   864: 'Spare_Fault_864', class No Acknowledgement, trigger "DB302_HMI_Faults_Carrier13_Faults_1" bit 15
   865: 'Carrier 13 Motion Off Fault', class No Acknowledgement, trigger "DB302_HMI_Faults_Carrier13_Faults_2" bit 0
   866: 'Carrier 13 Motion On Fault', class No Acknowledgement, trigger "DB302_HMI_Faults_Carrier13_Faults_2" bit 1
   867: 'Carrier 13 Spacing Fault', class No Acknowledgement, trigger "DB302_HMI_Faults_Carrier13_Faults_2" bit 2
   868: 'Carrier 13 Duplicate Carrier Number Fault', class No Acknowledgement, trigger "DB302_HMI_Faults_Carrier13_Faults_2" bit 3
   869: 'Spare_Fault_869', class No Acknowledgement, trigger "DB302_HMI_Faults_Carrier13_Faults_2" bit 4
   870: 'Spare_Fault_870', class No Acknowledgement, trigger "DB302_HMI_Faults_Carrier13_Faults_2" bit 5
   871: 'Spare_Fault_871', class No Acknowledgement, trigger "DB302_HMI_Faults_Carrier13_Faults_2" bit 6
   872: 'Spare_Fault_872', class No Acknowledgement, trigger "DB302_HMI_Faults_Carrier13_Faults_2" bit 7
   873: 'Spare_Fault_873', class No Acknowledgement, trigger "DB302_HMI_Faults_Carrier13_Faults_2" bit 8
   874: 'Spare_Fault_874', class No Acknowledgement, trigger "DB302_HMI_Faults_Carrier13_Faults_2" bit 9
   875: 'Spare_Fault_875', class No Acknowledgement, trigger "DB302_HMI_Faults_Carrier13_Faults_2" bit 10
   876: 'Spare_Fault_876', class No Acknowledgement, trigger "DB302_HMI_Faults_Carrier13_Faults_2" bit 11
   877: 'Spare_Fault_877', class No Acknowledgement, trigger "DB302_HMI_Faults_Carrier13_Faults_2" bit 12
   878: 'Spare_Fault_878', class No Acknowledgement, trigger "DB302_HMI_Faults_Carrier13_Faults_2" bit 13
   879: 'Spare_Fault_879', class No Acknowledgement, trigger "DB302_HMI_Faults_Carrier13_Faults_2" bit 14
   880: 'Spare_Fault_880', class No Acknowledgement, trigger "DB302_HMI_Faults_Carrier13_Faults_2" bit 15
   881: 'Spare_Fault_881', class No Acknowledgement, trigger "DB302_HMI_Faults_Carrier13_Faults_3" bit 0
   882: 'Spare_Fault_882', class No Acknowledgement, trigger "DB302_HMI_Faults_Carrier13_Faults_3" bit 1
   883: 'Spare_Fault_883', class No Acknowledgement, trigger "DB302_HMI_Faults_Carrier13_Faults_3" bit 2
   884: 'Spare_Fault_884', class No Acknowledgement, trigger "DB302_HMI_Faults_Carrier13_Faults_3" bit 3
   885: 'Spare_Fault_885', class No Acknowledgement, trigger "DB302_HMI_Faults_Carrier13_Faults_3" bit 4
   886: 'Spare_Fault_886', class No Acknowledgement, trigger "DB302_HMI_Faults_Carrier13_Faults_3" bit 5
   887: 'Spare_Fault_887', class No Acknowledgement, trigger "DB302_HMI_Faults_Carrier13_Faults_3" bit 6
   888: 'Spare_Fault_888', class No Acknowledgement, trigger "DB302_HMI_Faults_Carrier13_Faults_3" bit 7
   889: 'Spare_Fault_889', class No Acknowledgement, trigger "DB302_HMI_Faults_Carrier13_Faults_3" bit 8
   890: 'Spare_Fault_890', class No Acknowledgement, trigger "DB302_HMI_Faults_Carrier13_Faults_3" bit 9
   891: 'Spare_Fault_891', class No Acknowledgement, trigger "DB302_HMI_Faults_Carrier13_Faults_3" bit 10
   892: 'Spare_Fault_892', class No Acknowledgement, trigger "DB302_HMI_Faults_Carrier13_Faults_3" bit 11
   893: 'Spare_Fault_893', class No Acknowledgement, trigger "DB302_HMI_Faults_Carrier13_Faults_3" bit 12
   894: 'Spare_Fault_894', class No Acknowledgement, trigger "DB302_HMI_Faults_Carrier13_Faults_3" bit 13
   895: 'Spare_Fault_895', class No Acknowledgement, trigger "DB302_HMI_Faults_Carrier13_Faults_3" bit 14
   896: 'Spare_Fault_896', class No Acknowledgement, trigger "DB302_HMI_Faults_Carrier13_Faults_3" bit 15
   897: 'Carrier 14 Disconnect Open Power Fault DI11.0', class No Acknowledgement, trigger "DB302_HMI_Faults_Carrier14_Faults_0" bit 0
   898: 'Carrier 14 Drive Profinet Comm Fault', class No Acknowledgement, trigger "DB302_HMI_Faults_Carrier14_Faults_0" bit 1
   899: 'Carrier 14 Production Stop Not Reset', class No Acknowledgement, trigger "DB302_HMI_Faults_Carrier14_Faults_0" bit 2
   900: 'Carrier 14 CB02122 Tripped', class No Acknowledgement, trigger "DB302_HMI_Faults_Carrier14_Faults_0" bit 3
   901: 'Carrier 14 CB02123 Tripped', class No Acknowledgement, trigger "DB302_HMI_Faults_Carrier14_Faults_0" bit 4
   902: 'Carrier 14 AUX1 CB Tripped', class No Acknowledgement, trigger "DB302_HMI_Faults_Carrier14_Faults_0" bit 5
   903: 'Carrier 14 AUX2 CB Tripped', class No Acknowledgement, trigger "DB302_HMI_Faults_Carrier14_Faults_0" bit 6
   904: 'Carrier 14 PLC Not Communicating', class No Acknowledgement, trigger "DB302_HMI_Faults_Carrier14_Faults_0" bit 7
   905: 'Carrier 14 Safe Input Card Fault', class No Acknowledgement, trigger "DB302_HMI_Faults_Carrier14_Faults_0" bit 8
   906: 'Carrier 14 Safe Output Card Fault', class No Acknowledgement, trigger "DB302_HMI_Faults_Carrier14_Faults_0" bit 9
   907: 'Carrier 14 Standard Input Card Fault', class No Acknowledgement, trigger "DB302_HMI_Faults_Carrier14_Faults_0" bit 10
   908: 'Carrier 14 Standard Output Card Fault', class No Acknowledgement, trigger "DB302_HMI_Faults_Carrier14_Faults_0" bit 11
   909: 'Carrier 14 Encoder Position Fault', class No Acknowledgement, trigger "DB302_HMI_Faults_Carrier14_Faults_0" bit 12
   910: 'Carrier 14 Encoder Internal Error', class No Acknowledgement, trigger "DB302_HMI_Faults_Carrier14_Faults_0" bit 13
   911: 'Carrier 14 Encoder Comm Fault', class No Acknowledgement, trigger "DB302_HMI_Faults_Carrier14_Faults_0" bit 14
   912: 'Carrier 14 HMI Comm Fault', class No Acknowledgement, trigger "DB302_HMI_Faults_Carrier14_Faults_0" bit 15
   913: 'Carrier 14 Crash Detection Fault', class No Acknowledgement, trigger "DB302_HMI_Faults_Carrier14_Faults_1" bit 0
   914: 'Carrier 14 Carrier Number Invalid', class No Acknowledgement, trigger "DB302_HMI_Faults_Carrier14_Faults_1" bit 1
   915: 'Carrier 14 Drive: PROFINET configuration error', class No Acknowledgement, trigger "DB302_HMI_Faults_Carrier14_Faults_1" bit 2
   916: 'Carrier 14 Drive: Error internal communications', class No Acknowledgement, trigger "DB302_HMI_Faults_Carrier14_Faults_1" bit 3
   917: 'Carrier 14 Drive: Motor overtemperature', class No Acknowledgement, trigger "DB302_HMI_Faults_Carrier14_Faults_1" bit 4
   918: 'Carrier 14 Drive: Motor overcurrent', class No Acknowledgement, trigger "DB302_HMI_Faults_Carrier14_Faults_1" bit 5
   919: 'Carrier 14 Drive: Infeed or power unit not ready', class No Acknowledgement, trigger "DB302_HMI_Faults_Carrier14_Faults_1" bit 6
   920: 'Carrier 14 Drive: Short-circuit/ground fault detected', class No Acknowledgement, trigger "DB302_HMI_Faults_Carrier14_Faults_1" bit 7
   921: 'Carrier 14 Drive: PROFINET Setpoint timeout', class No Acknowledgement, trigger "DB302_HMI_Faults_Carrier14_Faults_1" bit 8
   922: 'Carrier 14 Power unit: Overcurrent', class No Acknowledgement, trigger "DB302_HMI_Faults_Carrier14_Faults_1" bit 9
   923: 'Carrier 14 Power unit: DC link voltage overvoltage', class No Acknowledgement, trigger "DB302_HMI_Faults_Carrier14_Faults_1" bit 10
   924: 'Carrier 14 Power unit: DC link voltage undervoltage', class No Acknowledgement, trigger "DB302_HMI_Faults_Carrier14_Faults_1" bit 11
   925: 'Carrier 14 Power unit: Line phase failure in main circuit', class No Acknowledgement, trigger "DB302_HMI_Faults_Carrier14_Faults_1" bit 12
   926: 'Carrier 14 Power unit: Phase failure motor cable', class No Acknowledgement, trigger "DB302_HMI_Faults_Carrier14_Faults_1" bit 13
   927: 'Carrier 14 Power unit: Ground fault', class No Acknowledgement, trigger "DB302_HMI_Faults_Carrier14_Faults_1" bit 14
   928: 'Spare_Fault_928', class No Acknowledgement, trigger "DB302_HMI_Faults_Carrier14_Faults_1" bit 15
   929: 'Carrier 14 Motion Off Fault', class No Acknowledgement, trigger "DB302_HMI_Faults_Carrier14_Faults_2" bit 0
   930: 'Carrier 14 Motion On Fault', class No Acknowledgement, trigger "DB302_HMI_Faults_Carrier14_Faults_2" bit 1
   931: 'Carrier 14 Spacing Fault', class No Acknowledgement, trigger "DB302_HMI_Faults_Carrier14_Faults_2" bit 2
   932: 'Carrier 14 Duplicate Carrier Number Fault', class No Acknowledgement, trigger "DB302_HMI_Faults_Carrier14_Faults_2" bit 3
   933: 'Spare_Fault_933', class No Acknowledgement, trigger "DB302_HMI_Faults_Carrier14_Faults_2" bit 4
   934: 'Spare_Fault_934', class No Acknowledgement, trigger "DB302_HMI_Faults_Carrier14_Faults_2" bit 5
   935: 'Spare_Fault_935', class No Acknowledgement, trigger "DB302_HMI_Faults_Carrier14_Faults_2" bit 6
   936: 'Spare_Fault_936', class No Acknowledgement, trigger "DB302_HMI_Faults_Carrier14_Faults_2" bit 7
   937: 'Spare_Fault_937', class No Acknowledgement, trigger "DB302_HMI_Faults_Carrier14_Faults_2" bit 8
   938: 'Spare_Fault_938', class No Acknowledgement, trigger "DB302_HMI_Faults_Carrier14_Faults_2" bit 9
   939: 'Spare_Fault_939', class No Acknowledgement, trigger "DB302_HMI_Faults_Carrier14_Faults_2" bit 10
   940: 'Spare_Fault_940', class No Acknowledgement, trigger "DB302_HMI_Faults_Carrier14_Faults_2" bit 11
   941: 'Spare_Fault_941', class No Acknowledgement, trigger "DB302_HMI_Faults_Carrier14_Faults_2" bit 12
   942: 'Spare_Fault_942', class No Acknowledgement, trigger "DB302_HMI_Faults_Carrier14_Faults_2" bit 13
   943: 'Spare_Fault_943', class No Acknowledgement, trigger "DB302_HMI_Faults_Carrier14_Faults_2" bit 14
   944: 'Spare_Fault_944', class No Acknowledgement, trigger "DB302_HMI_Faults_Carrier14_Faults_2" bit 15
   945: 'Spare_Fault_945', class No Acknowledgement, trigger "DB302_HMI_Faults_Carrier14_Faults_3" bit 0
   946: 'Spare_Fault_946', class No Acknowledgement, trigger "DB302_HMI_Faults_Carrier14_Faults_3" bit 1
   947: 'Spare_Fault_947', class No Acknowledgement, trigger "DB302_HMI_Faults_Carrier14_Faults_3" bit 2
   948: 'Spare_Fault_948', class No Acknowledgement, trigger "DB302_HMI_Faults_Carrier14_Faults_3" bit 3
   949: 'Spare_Fault_949', class No Acknowledgement, trigger "DB302_HMI_Faults_Carrier14_Faults_3" bit 4
   950: 'Spare_Fault_950', class No Acknowledgement, trigger "DB302_HMI_Faults_Carrier14_Faults_3" bit 5
   951: 'Spare_Fault_951', class No Acknowledgement, trigger "DB302_HMI_Faults_Carrier14_Faults_3" bit 6
   952: 'Spare_Fault_952', class No Acknowledgement, trigger "DB302_HMI_Faults_Carrier14_Faults_3" bit 7
   953: 'Spare_Fault_953', class No Acknowledgement, trigger "DB302_HMI_Faults_Carrier14_Faults_3" bit 8
   954: 'Spare_Fault_954', class No Acknowledgement, trigger "DB302_HMI_Faults_Carrier14_Faults_3" bit 9
   955: 'Spare_Fault_955', class No Acknowledgement, trigger "DB302_HMI_Faults_Carrier14_Faults_3" bit 10
   956: 'Spare_Fault_956', class No Acknowledgement, trigger "DB302_HMI_Faults_Carrier14_Faults_3" bit 11
   957: 'Spare_Fault_957', class No Acknowledgement, trigger "DB302_HMI_Faults_Carrier14_Faults_3" bit 12
   958: 'Spare_Fault_958', class No Acknowledgement, trigger "DB302_HMI_Faults_Carrier14_Faults_3" bit 13
   959: 'Spare_Fault_959', class No Acknowledgement, trigger "DB302_HMI_Faults_Carrier14_Faults_3" bit 14
   960: 'Spare_Fault_960', class No Acknowledgement, trigger "DB302_HMI_Faults_Carrier14_Faults_3" bit 15
   961: 'Carrier 15 Disconnect Open Power Fault DI11.0', class No Acknowledgement, trigger "DB302_HMI_Faults_Carrier15_Faults_0" bit 0
   962: 'Carrier 15 Drive Profinet Comm Fault', class No Acknowledgement, trigger "DB302_HMI_Faults_Carrier15_Faults_0" bit 1
   963: 'Carrier 15 Production Stop Not Reset', class No Acknowledgement, trigger "DB302_HMI_Faults_Carrier15_Faults_0" bit 2
   964: 'Carrier 15 CB02122 Tripped', class No Acknowledgement, trigger "DB302_HMI_Faults_Carrier15_Faults_0" bit 3
   965: 'Carrier 15 CB02123 Tripped', class No Acknowledgement, trigger "DB302_HMI_Faults_Carrier15_Faults_0" bit 4
   966: 'Carrier 15 AUX1 CB Tripped', class No Acknowledgement, trigger "DB302_HMI_Faults_Carrier15_Faults_0" bit 5
   967: 'Carrier 15 AUX2 CB Tripped', class No Acknowledgement, trigger "DB302_HMI_Faults_Carrier15_Faults_0" bit 6
   968: 'Carrier 15 PLC Not Communicating', class No Acknowledgement, trigger "DB302_HMI_Faults_Carrier15_Faults_0" bit 7
   969: 'Carrier 15 Safe Input Card Fault', class No Acknowledgement, trigger "DB302_HMI_Faults_Carrier15_Faults_0" bit 8
   970: 'Carrier 15 Safe Output Card Fault', class No Acknowledgement, trigger "DB302_HMI_Faults_Carrier15_Faults_0" bit 9
   971: 'Carrier 15 Standard Input Card Fault', class No Acknowledgement, trigger "DB302_HMI_Faults_Carrier15_Faults_0" bit 10
   972: 'Carrier 15 Standard Output Card Fault', class No Acknowledgement, trigger "DB302_HMI_Faults_Carrier15_Faults_0" bit 11
   973: 'Carrier 15 Encoder Position Fault', class No Acknowledgement, trigger "DB302_HMI_Faults_Carrier15_Faults_0" bit 12
   974: 'Carrier 15 Encoder Internal Error', class No Acknowledgement, trigger "DB302_HMI_Faults_Carrier15_Faults_0" bit 13
   975: 'Carrier 15 Encoder Comm Fault', class No Acknowledgement, trigger "DB302_HMI_Faults_Carrier15_Faults_0" bit 14
   976: 'Carrier 15 HMI Comm Fault', class No Acknowledgement, trigger "DB302_HMI_Faults_Carrier15_Faults_0" bit 15
   977: 'Carrier 15 Crash Detection Fault', class No Acknowledgement, trigger "DB302_HMI_Faults_Carrier15_Faults_1" bit 0
   978: 'Carrier 15 Carrier Number Invalid', class No Acknowledgement, trigger "DB302_HMI_Faults_Carrier15_Faults_1" bit 1
   979: 'Carrier 15 Drive: PROFINET configuration error', class No Acknowledgement, trigger "DB302_HMI_Faults_Carrier15_Faults_1" bit 2
   980: 'Carrier 15 Drive: Error internal communications', class No Acknowledgement, trigger "DB302_HMI_Faults_Carrier15_Faults_1" bit 3
   981: 'Carrier 15 Drive: Motor overtemperature', class No Acknowledgement, trigger "DB302_HMI_Faults_Carrier15_Faults_1" bit 4
   982: 'Carrier 15 Drive: Motor overcurrent', class No Acknowledgement, trigger "DB302_HMI_Faults_Carrier15_Faults_1" bit 5
   983: 'Carrier 15 Drive: Infeed or power unit not ready', class No Acknowledgement, trigger "DB302_HMI_Faults_Carrier15_Faults_1" bit 6
   984: 'Carrier 15 Drive: Short-circuit/ground fault detected', class No Acknowledgement, trigger "DB302_HMI_Faults_Carrier15_Faults_1" bit 7
   985: 'Carrier 15 Drive: PROFINET Setpoint timeout', class No Acknowledgement, trigger "DB302_HMI_Faults_Carrier15_Faults_1" bit 8
   986: 'Carrier 15 Power unit: Overcurrent', class No Acknowledgement, trigger "DB302_HMI_Faults_Carrier15_Faults_1" bit 9
   987: 'Carrier 15 Power unit: DC link voltage overvoltage', class No Acknowledgement, trigger "DB302_HMI_Faults_Carrier15_Faults_1" bit 10
   988: 'Carrier 15 Power unit: DC link voltage undervoltage', class No Acknowledgement, trigger "DB302_HMI_Faults_Carrier15_Faults_1" bit 11
   989: 'Carrier 15 Power unit: Line phase failure in main circuit', class No Acknowledgement, trigger "DB302_HMI_Faults_Carrier15_Faults_1" bit 12
   990: 'Carrier 15 Power unit: Phase failure motor cable', class No Acknowledgement, trigger "DB302_HMI_Faults_Carrier15_Faults_1" bit 13
   991: 'Carrier 15 Power unit: Ground fault', class No Acknowledgement, trigger "DB302_HMI_Faults_Carrier15_Faults_1" bit 14
   992: 'Spare_Fault_992', class No Acknowledgement, trigger "DB302_HMI_Faults_Carrier15_Faults_1" bit 15
   993: 'Carrier 15 Motion Off Fault', class No Acknowledgement, trigger "DB302_HMI_Faults_Carrier15_Faults_2" bit 0
   994: 'Carrier 15 Motion On Fault', class No Acknowledgement, trigger "DB302_HMI_Faults_Carrier15_Faults_2" bit 1
   995: 'Carrier 15 Spacing Fault', class No Acknowledgement, trigger "DB302_HMI_Faults_Carrier15_Faults_2" bit 2
   996: 'Carrier 15 Duplicate Carrier Number Fault', class No Acknowledgement, trigger "DB302_HMI_Faults_Carrier15_Faults_2" bit 3
   997: 'Spare_Fault_997', class No Acknowledgement, trigger "DB302_HMI_Faults_Carrier15_Faults_2" bit 4
   998: 'Spare_Fault_998', class No Acknowledgement, trigger "DB302_HMI_Faults_Carrier15_Faults_2" bit 5
   999: 'Spare_Fault_999', class No Acknowledgement, trigger "DB302_HMI_Faults_Carrier15_Faults_2" bit 6
   1000: 'Spare_Fault_1000', class No Acknowledgement, trigger "DB302_HMI_Faults_Carrier15_Faults_2" bit 7
   1001: 'Spare_Fault_1001', class No Acknowledgement, trigger "DB302_HMI_Faults_Carrier15_Faults_2" bit 8
   1002: 'Spare_Fault_1002', class No Acknowledgement, trigger "DB302_HMI_Faults_Carrier15_Faults_2" bit 9
   1003: 'Spare_Fault_1003', class No Acknowledgement, trigger "DB302_HMI_Faults_Carrier15_Faults_2" bit 10
   1004: 'Spare_Fault_1004', class No Acknowledgement, trigger "DB302_HMI_Faults_Carrier15_Faults_2" bit 11
   1005: 'Spare_Fault_1005', class No Acknowledgement, trigger "DB302_HMI_Faults_Carrier15_Faults_2" bit 12
   1006: 'Spare_Fault_1006', class No Acknowledgement, trigger "DB302_HMI_Faults_Carrier15_Faults_2" bit 13
   1007: 'Spare_Fault_1007', class No Acknowledgement, trigger "DB302_HMI_Faults_Carrier15_Faults_2" bit 14
   1008: 'Spare_Fault_1008', class No Acknowledgement, trigger "DB302_HMI_Faults_Carrier15_Faults_2" bit 15
   1009: 'Spare_Fault_1009', class No Acknowledgement, trigger "DB302_HMI_Faults_Carrier15_Faults_3" bit 0
   1010: 'Spare_Fault_1010', class No Acknowledgement, trigger "DB302_HMI_Faults_Carrier15_Faults_3" bit 1
   1011: 'Spare_Fault_1011', class No Acknowledgement, trigger "DB302_HMI_Faults_Carrier15_Faults_3" bit 2
   1012: 'Spare_Fault_1012', class No Acknowledgement, trigger "DB302_HMI_Faults_Carrier15_Faults_3" bit 3
   1013: 'Spare_Fault_1013', class No Acknowledgement, trigger "DB302_HMI_Faults_Carrier15_Faults_3" bit 4
   1014: 'Spare_Fault_1014', class No Acknowledgement, trigger "DB302_HMI_Faults_Carrier15_Faults_3" bit 5
   1015: 'Spare_Fault_1015', class No Acknowledgement, trigger "DB302_HMI_Faults_Carrier15_Faults_3" bit 6
   1016: 'Spare_Fault_1016', class No Acknowledgement, trigger "DB302_HMI_Faults_Carrier15_Faults_3" bit 7
   1017: 'Spare_Fault_1017', class No Acknowledgement, trigger "DB302_HMI_Faults_Carrier15_Faults_3" bit 8
   1018: 'Spare_Fault_1018', class No Acknowledgement, trigger "DB302_HMI_Faults_Carrier15_Faults_3" bit 9
   1019: 'Spare_Fault_1019', class No Acknowledgement, trigger "DB302_HMI_Faults_Carrier15_Faults_3" bit 10
   1020: 'Spare_Fault_1020', class No Acknowledgement, trigger "DB302_HMI_Faults_Carrier15_Faults_3" bit 11
   1021: 'Spare_Fault_1021', class No Acknowledgement, trigger "DB302_HMI_Faults_Carrier15_Faults_3" bit 12
   1022: 'Spare_Fault_1022', class No Acknowledgement, trigger "DB302_HMI_Faults_Carrier15_Faults_3" bit 13
   1023: 'Spare_Fault_1023', class No Acknowledgement, trigger "DB302_HMI_Faults_Carrier15_Faults_3" bit 14
   1024: 'Spare_Fault_1024', class No Acknowledgement, trigger "DB302_HMI_Faults_Carrier15_Faults_3" bit 15
   1025: 'Carrier 16 Disconnect Open Power Fault DI11.0', class No Acknowledgement, trigger "DB302_HMI_Faults_Carrier16_Faults_0" bit 0
   1026: 'Carrier 16 Drive Profinet Comm Fault', class No Acknowledgement, trigger "DB302_HMI_Faults_Carrier16_Faults_0" bit 1
   1027: 'Carrier 16 Production Stop Not Reset', class No Acknowledgement, trigger "DB302_HMI_Faults_Carrier16_Faults_0" bit 2
   1028: 'Carrier 16 CB02122 Tripped', class No Acknowledgement, trigger "DB302_HMI_Faults_Carrier16_Faults_0" bit 3
   1029: 'Carrier 16 CB02123 Tripped', class No Acknowledgement, trigger "DB302_HMI_Faults_Carrier16_Faults_0" bit 4
   1030: 'Carrier 16 AUX1 CB Tripped', class No Acknowledgement, trigger "DB302_HMI_Faults_Carrier16_Faults_0" bit 5
   1031: 'Carrier 16 AUX2 CB Tripped', class No Acknowledgement, trigger "DB302_HMI_Faults_Carrier16_Faults_0" bit 6
   1032: 'Carrier 16 PLC Not Communicating', class No Acknowledgement, trigger "DB302_HMI_Faults_Carrier16_Faults_0" bit 7
   1033: 'Carrier 16 Safe Input Card Fault', class No Acknowledgement, trigger "DB302_HMI_Faults_Carrier16_Faults_0" bit 8
   1034: 'Carrier 16 Safe Output Card Fault', class No Acknowledgement, trigger "DB302_HMI_Faults_Carrier16_Faults_0" bit 9
   1035: 'Carrier 16 Standard Input Card Fault', class No Acknowledgement, trigger "DB302_HMI_Faults_Carrier16_Faults_0" bit 10
   1036: 'Carrier 16 Standard Output Card Fault', class No Acknowledgement, trigger "DB302_HMI_Faults_Carrier16_Faults_0" bit 11
   1037: 'Carrier 16 Encoder Position Fault', class No Acknowledgement, trigger "DB302_HMI_Faults_Carrier16_Faults_0" bit 12
   1038: 'Carrier 16 Encoder Internal Error', class No Acknowledgement, trigger "DB302_HMI_Faults_Carrier16_Faults_0" bit 13
   1039: 'Carrier 16 Encoder Comm Fault', class No Acknowledgement, trigger "DB302_HMI_Faults_Carrier16_Faults_0" bit 14
   1040: 'Carrier 16 HMI Comm Fault', class No Acknowledgement, trigger "DB302_HMI_Faults_Carrier16_Faults_0" bit 15
   1041: 'Carrier 16 Crash Detection Fault', class No Acknowledgement, trigger "DB302_HMI_Faults_Carrier16_Faults_1" bit 0
   1042: 'Carrier 16 Carrier Number Invalid', class No Acknowledgement, trigger "DB302_HMI_Faults_Carrier16_Faults_1" bit 1
   1043: 'Carrier 16 Drive: PROFINET configuration error', class No Acknowledgement, trigger "DB302_HMI_Faults_Carrier16_Faults_1" bit 2
   1044: 'Carrier 16 Drive: Error internal communications', class No Acknowledgement, trigger "DB302_HMI_Faults_Carrier16_Faults_1" bit 3
   1045: 'Carrier 16 Drive: Motor overtemperature', class No Acknowledgement, trigger "DB302_HMI_Faults_Carrier16_Faults_1" bit 4
   1046: 'Carrier 16 Drive: Motor overcurrent', class No Acknowledgement, trigger "DB302_HMI_Faults_Carrier16_Faults_1" bit 5
   1047: 'Carrier 16 Drive: Infeed or power unit not ready', class No Acknowledgement, trigger "DB302_HMI_Faults_Carrier16_Faults_1" bit 6
   1048: 'Carrier 16 Drive: Short-circuit/ground fault detected', class No Acknowledgement, trigger "DB302_HMI_Faults_Carrier16_Faults_1" bit 7
   1049: 'Carrier 16 Drive: PROFINET Setpoint timeout', class No Acknowledgement, trigger "DB302_HMI_Faults_Carrier16_Faults_1" bit 8
   1050: 'Carrier 16 Power unit: Overcurrent', class No Acknowledgement, trigger "DB302_HMI_Faults_Carrier16_Faults_1" bit 9
   1051: 'Carrier 16 Power unit: DC link voltage overvoltage', class No Acknowledgement, trigger "DB302_HMI_Faults_Carrier16_Faults_1" bit 10
   1052: 'Carrier 16 Power unit: DC link voltage undervoltage', class No Acknowledgement, trigger "DB302_HMI_Faults_Carrier16_Faults_1" bit 11
   1053: 'Carrier 16 Power unit: Line phase failure in main circuit', class No Acknowledgement, trigger "DB302_HMI_Faults_Carrier16_Faults_1" bit 12
   1054: 'Carrier 16 Power unit: Phase failure motor cable', class No Acknowledgement, trigger "DB302_HMI_Faults_Carrier16_Faults_1" bit 13
   1055: 'Carrier 16 Power unit: Ground fault', class No Acknowledgement, trigger "DB302_HMI_Faults_Carrier16_Faults_1" bit 14
   1056: 'Spare_Fault_1056', class No Acknowledgement, trigger "DB302_HMI_Faults_Carrier16_Faults_1" bit 15
   1057: 'Carrier 16 Motion Off Fault', class No Acknowledgement, trigger "DB302_HMI_Faults_Carrier16_Faults_2" bit 0
   1058: 'Carrier 16 Motion On Fault', class No Acknowledgement, trigger "DB302_HMI_Faults_Carrier16_Faults_2" bit 1
   1059: 'Carrier 16 Spacing Fault', class No Acknowledgement, trigger "DB302_HMI_Faults_Carrier16_Faults_2" bit 2
   1060: 'Carrier 16 Duplicate Carrier Number Fault', class No Acknowledgement, trigger "DB302_HMI_Faults_Carrier16_Faults_2" bit 3
   1061: 'Spare_Fault_1061', class No Acknowledgement, trigger "DB302_HMI_Faults_Carrier16_Faults_2" bit 4
   1062: 'Spare_Fault_1062', class No Acknowledgement, trigger "DB302_HMI_Faults_Carrier16_Faults_2" bit 5
   1063: 'Spare_Fault_1063', class No Acknowledgement, trigger "DB302_HMI_Faults_Carrier16_Faults_2" bit 6
   1064: 'Spare_Fault_1064', class No Acknowledgement, trigger "DB302_HMI_Faults_Carrier16_Faults_2" bit 7
   1065: 'Spare_Fault_1065', class No Acknowledgement, trigger "DB302_HMI_Faults_Carrier16_Faults_2" bit 8
   1066: 'Spare_Fault_1066', class No Acknowledgement, trigger "DB302_HMI_Faults_Carrier16_Faults_2" bit 9
   1067: 'Spare_Fault_1067', class No Acknowledgement, trigger "DB302_HMI_Faults_Carrier16_Faults_2" bit 10
   1068: 'Spare_Fault_1068', class No Acknowledgement, trigger "DB302_HMI_Faults_Carrier16_Faults_2" bit 11
   1069: 'Spare_Fault_1069', class No Acknowledgement, trigger "DB302_HMI_Faults_Carrier16_Faults_2" bit 12
   1070: 'Spare_Fault_1070', class No Acknowledgement, trigger "DB302_HMI_Faults_Carrier16_Faults_2" bit 13
   1071: 'Spare_Fault_1071', class No Acknowledgement, trigger "DB302_HMI_Faults_Carrier16_Faults_2" bit 14
   1072: 'Spare_Fault_1072', class No Acknowledgement, trigger "DB302_HMI_Faults_Carrier16_Faults_2" bit 15
   1073: 'Spare_Fault_1073', class No Acknowledgement, trigger "DB302_HMI_Faults_Carrier16_Faults_3" bit 0
   1074: 'Spare_Fault_1074', class No Acknowledgement, trigger "DB302_HMI_Faults_Carrier16_Faults_3" bit 1
   1075: 'Spare_Fault_1075', class No Acknowledgement, trigger "DB302_HMI_Faults_Carrier16_Faults_3" bit 2
   1076: 'Spare_Fault_1076', class No Acknowledgement, trigger "DB302_HMI_Faults_Carrier16_Faults_3" bit 3
   1077: 'Spare_Fault_1077', class No Acknowledgement, trigger "DB302_HMI_Faults_Carrier16_Faults_3" bit 4
   1078: 'Spare_Fault_1078', class No Acknowledgement, trigger "DB302_HMI_Faults_Carrier16_Faults_3" bit 5
   1079: 'Spare_Fault_1079', class No Acknowledgement, trigger "DB302_HMI_Faults_Carrier16_Faults_3" bit 6
   1080: 'Spare_Fault_1080', class No Acknowledgement, trigger "DB302_HMI_Faults_Carrier16_Faults_3" bit 7
   1081: 'Spare_Fault_1081', class No Acknowledgement, trigger "DB302_HMI_Faults_Carrier16_Faults_3" bit 8
   1082: 'Spare_Fault_1082', class No Acknowledgement, trigger "DB302_HMI_Faults_Carrier16_Faults_3" bit 9
   1083: 'Spare_Fault_1083', class No Acknowledgement, trigger "DB302_HMI_Faults_Carrier16_Faults_3" bit 10
   1084: 'Spare_Fault_1084', class No Acknowledgement, trigger "DB302_HMI_Faults_Carrier16_Faults_3" bit 11
   1085: 'Spare_Fault_1085', class No Acknowledgement, trigger "DB302_HMI_Faults_Carrier16_Faults_3" bit 12
   1086: 'Spare_Fault_1086', class No Acknowledgement, trigger "DB302_HMI_Faults_Carrier16_Faults_3" bit 13
   1087: 'Spare_Fault_1087', class No Acknowledgement, trigger "DB302_HMI_Faults_Carrier16_Faults_3" bit 14
   1088: 'Spare_Fault_1088', class No Acknowledgement, trigger "DB302_HMI_Faults_Carrier16_Faults_3" bit 15
   1089: 'Carrier 17 Disconnect Open Power Fault DI11.0', class No Acknowledgement, trigger "DB302_HMI_Faults_Carrier17_Faults_0" bit 0
   1090: 'Carrier 17 Drive Profinet Comm Fault', class No Acknowledgement, trigger "DB302_HMI_Faults_Carrier17_Faults_0" bit 1
   1091: 'Carrier 17 Production Stop Not Reset', class No Acknowledgement, trigger "DB302_HMI_Faults_Carrier17_Faults_0" bit 2
   1092: 'Carrier 17 CB02122 Tripped', class No Acknowledgement, trigger "DB302_HMI_Faults_Carrier17_Faults_0" bit 3
   1093: 'Carrier 17 CB02123 Tripped', class No Acknowledgement, trigger "DB302_HMI_Faults_Carrier17_Faults_0" bit 4
   1094: 'Carrier 17 AUX1 CB Tripped', class No Acknowledgement, trigger "DB302_HMI_Faults_Carrier17_Faults_0" bit 5
   1095: 'Carrier 17 AUX2 CB Tripped', class No Acknowledgement, trigger "DB302_HMI_Faults_Carrier17_Faults_0" bit 6
   1096: 'Carrier 17 PLC Not Communicating', class No Acknowledgement, trigger "DB302_HMI_Faults_Carrier17_Faults_0" bit 7
   1097: 'Carrier 17 Safe Input Card Fault', class No Acknowledgement, trigger "DB302_HMI_Faults_Carrier17_Faults_0" bit 8
   1098: 'Carrier 17 Safe Output Card Fault', class No Acknowledgement, trigger "DB302_HMI_Faults_Carrier17_Faults_0" bit 9
   1099: 'Carrier 17 Standard Input Card Fault', class No Acknowledgement, trigger "DB302_HMI_Faults_Carrier17_Faults_0" bit 10
   1100: 'Carrier 17 Standard Output Card Fault', class No Acknowledgement, trigger "DB302_HMI_Faults_Carrier17_Faults_0" bit 11
   1101: 'Carrier 17 Encoder Position Fault', class No Acknowledgement, trigger "DB302_HMI_Faults_Carrier17_Faults_0" bit 12
   1102: 'Carrier 17 Encoder Internal Error', class No Acknowledgement, trigger "DB302_HMI_Faults_Carrier17_Faults_0" bit 13
   1103: 'Carrier 17 Encoder Comm Fault', class No Acknowledgement, trigger "DB302_HMI_Faults_Carrier17_Faults_0" bit 14
   1104: 'Carrier 17 HMI Comm Fault', class No Acknowledgement, trigger "DB302_HMI_Faults_Carrier17_Faults_0" bit 15
   1105: 'Carrier 17 Crash Detection Fault', class No Acknowledgement, trigger "DB302_HMI_Faults_Carrier17_Faults_1" bit 0
   1106: 'Carrier 17 Carrier Number Invalid', class No Acknowledgement, trigger "DB302_HMI_Faults_Carrier17_Faults_1" bit 1
   1107: 'Carrier 17 Drive: PROFINET configuration error', class No Acknowledgement, trigger "DB302_HMI_Faults_Carrier17_Faults_1" bit 2
   1108: 'Carrier 17 Drive: Error internal communications', class No Acknowledgement, trigger "DB302_HMI_Faults_Carrier17_Faults_1" bit 3
   1109: 'Carrier 17 Drive: Motor overtemperature', class No Acknowledgement, trigger "DB302_HMI_Faults_Carrier17_Faults_1" bit 4
   1110: 'Carrier 17 Drive: Motor overcurrent', class No Acknowledgement, trigger "DB302_HMI_Faults_Carrier17_Faults_1" bit 5
   1111: 'Carrier 17 Drive: Infeed or power unit not ready', class No Acknowledgement, trigger "DB302_HMI_Faults_Carrier17_Faults_1" bit 6
   1112: 'Carrier 17 Drive: Short-circuit/ground fault detected', class No Acknowledgement, trigger "DB302_HMI_Faults_Carrier17_Faults_1" bit 7
   1113: 'Carrier 17 Drive: PROFINET Setpoint timeout', class No Acknowledgement, trigger "DB302_HMI_Faults_Carrier17_Faults_1" bit 8
   1114: 'Carrier 17 Power unit: Overcurrent', class No Acknowledgement, trigger "DB302_HMI_Faults_Carrier17_Faults_1" bit 9
   1115: 'Carrier 17 Power unit: DC link voltage overvoltage', class No Acknowledgement, trigger "DB302_HMI_Faults_Carrier17_Faults_1" bit 10
   1116: 'Carrier 17 Power unit: DC link voltage undervoltage', class No Acknowledgement, trigger "DB302_HMI_Faults_Carrier17_Faults_1" bit 11
   1117: 'Carrier 17 Power unit: Line phase failure in main circuit', class No Acknowledgement, trigger "DB302_HMI_Faults_Carrier17_Faults_1" bit 12
   1118: 'Carrier 17 Power unit: Phase failure motor cable', class No Acknowledgement, trigger "DB302_HMI_Faults_Carrier17_Faults_1" bit 13
   1119: 'Carrier 17 Power unit: Ground fault', class No Acknowledgement, trigger "DB302_HMI_Faults_Carrier17_Faults_1" bit 14
   1120: 'Spare_Fault_1120', class No Acknowledgement, trigger "DB302_HMI_Faults_Carrier17_Faults_1" bit 15
   1121: 'Carrier 17 Motion Off Fault', class No Acknowledgement, trigger "DB302_HMI_Faults_Carrier17_Faults_2" bit 0
   1122: 'Carrier 17 Motion On Fault', class No Acknowledgement, trigger "DB302_HMI_Faults_Carrier17_Faults_2" bit 1
   1123: 'Carrier 17 Spacing Fault', class No Acknowledgement, trigger "DB302_HMI_Faults_Carrier17_Faults_2" bit 2
   1124: 'Carrier 17 Duplicate Carrier Number Fault', class No Acknowledgement, trigger "DB302_HMI_Faults_Carrier17_Faults_2" bit 3
   1125: 'Spare_Fault_1125', class No Acknowledgement, trigger "DB302_HMI_Faults_Carrier17_Faults_2" bit 4
   1126: 'Spare_Fault_1126', class No Acknowledgement, trigger "DB302_HMI_Faults_Carrier17_Faults_2" bit 5
   1127: 'Spare_Fault_1127', class No Acknowledgement, trigger "DB302_HMI_Faults_Carrier17_Faults_2" bit 6
   1128: 'Spare_Fault_1128', class No Acknowledgement, trigger "DB302_HMI_Faults_Carrier17_Faults_2" bit 7
   1129: 'Spare_Fault_1129', class No Acknowledgement, trigger "DB302_HMI_Faults_Carrier17_Faults_2" bit 8
   1130: 'Spare_Fault_1130', class No Acknowledgement, trigger "DB302_HMI_Faults_Carrier17_Faults_2" bit 9
   1131: 'Spare_Fault_1131', class No Acknowledgement, trigger "DB302_HMI_Faults_Carrier17_Faults_2" bit 10
   1132: 'Spare_Fault_1132', class No Acknowledgement, trigger "DB302_HMI_Faults_Carrier17_Faults_2" bit 11
   1133: 'Spare_Fault_1133', class No Acknowledgement, trigger "DB302_HMI_Faults_Carrier17_Faults_2" bit 12
   1134: 'Spare_Fault_1134', class No Acknowledgement, trigger "DB302_HMI_Faults_Carrier17_Faults_2" bit 13
   1135: 'Spare_Fault_1135', class No Acknowledgement, trigger "DB302_HMI_Faults_Carrier17_Faults_2" bit 14
   1136: 'Spare_Fault_1136', class No Acknowledgement, trigger "DB302_HMI_Faults_Carrier17_Faults_2" bit 15
   1137: 'Spare_Fault_1137', class No Acknowledgement, trigger "DB302_HMI_Faults_Carrier17_Faults_3" bit 0
   1138: 'Spare_Fault_1138', class No Acknowledgement, trigger "DB302_HMI_Faults_Carrier17_Faults_3" bit 1
   1139: 'Spare_Fault_1139', class No Acknowledgement, trigger "DB302_HMI_Faults_Carrier17_Faults_3" bit 2
   1140: 'Spare_Fault_1140', class No Acknowledgement, trigger "DB302_HMI_Faults_Carrier17_Faults_3" bit 3
   1141: 'Spare_Fault_1141', class No Acknowledgement, trigger "DB302_HMI_Faults_Carrier17_Faults_3" bit 4
   1142: 'Spare_Fault_1142', class No Acknowledgement, trigger "DB302_HMI_Faults_Carrier17_Faults_3" bit 5
   1143: 'Spare_Fault_1143', class No Acknowledgement, trigger "DB302_HMI_Faults_Carrier17_Faults_3" bit 6
   1144: 'Spare_Fault_1144', class No Acknowledgement, trigger "DB302_HMI_Faults_Carrier17_Faults_3" bit 7
   1145: 'Spare_Fault_1145', class No Acknowledgement, trigger "DB302_HMI_Faults_Carrier17_Faults_3" bit 8
   1146: 'Spare_Fault_1146', class No Acknowledgement, trigger "DB302_HMI_Faults_Carrier17_Faults_3" bit 9
   1147: 'Spare_Fault_1147', class No Acknowledgement, trigger "DB302_HMI_Faults_Carrier17_Faults_3" bit 10
   1148: 'Spare_Fault_1148', class No Acknowledgement, trigger "DB302_HMI_Faults_Carrier17_Faults_3" bit 11
   1149: 'Spare_Fault_1149', class No Acknowledgement, trigger "DB302_HMI_Faults_Carrier17_Faults_3" bit 12
   1150: 'Spare_Fault_1150', class No Acknowledgement, trigger "DB302_HMI_Faults_Carrier17_Faults_3" bit 13
   1151: 'Spare_Fault_1151', class No Acknowledgement, trigger "DB302_HMI_Faults_Carrier17_Faults_3" bit 14
   1152: 'Spare_Fault_1152', class No Acknowledgement, trigger "DB302_HMI_Faults_Carrier17_Faults_3" bit 15
   1153: 'Carrier 18 Disconnect Open Power Fault DI11.0', class No Acknowledgement, trigger "DB302_HMI_Faults_Carrier18_Faults_0" bit 0
   1154: 'Carrier 18 Drive Profinet Comm Fault', class No Acknowledgement, trigger "DB302_HMI_Faults_Carrier18_Faults_0" bit 1
   1155: 'Carrier 18 Production Stop Not Reset', class No Acknowledgement, trigger "DB302_HMI_Faults_Carrier18_Faults_0" bit 2
   1156: 'Carrier 18 CB02122 Tripped', class No Acknowledgement, trigger "DB302_HMI_Faults_Carrier18_Faults_0" bit 3
   1157: 'Carrier 18 CB02123 Tripped', class No Acknowledgement, trigger "DB302_HMI_Faults_Carrier18_Faults_0" bit 4
   1158: 'Carrier 18 AUX1 CB Tripped', class No Acknowledgement, trigger "DB302_HMI_Faults_Carrier18_Faults_0" bit 5
   1159: 'Carrier 18 AUX2 CB Tripped', class No Acknowledgement, trigger "DB302_HMI_Faults_Carrier18_Faults_0" bit 6
   1160: 'Carrier 18 PLC Not Communicating', class No Acknowledgement, trigger "DB302_HMI_Faults_Carrier18_Faults_0" bit 7
   1161: 'Carrier 18 Safe Input Card Fault', class No Acknowledgement, trigger "DB302_HMI_Faults_Carrier18_Faults_0" bit 8
   1162: 'Carrier 18 Safe Output Card Fault', class No Acknowledgement, trigger "DB302_HMI_Faults_Carrier18_Faults_0" bit 9
   1163: 'Carrier 18 Standard Input Card Fault', class No Acknowledgement, trigger "DB302_HMI_Faults_Carrier18_Faults_0" bit 10
   1164: 'Carrier 18 Standard Output Card Fault', class No Acknowledgement, trigger "DB302_HMI_Faults_Carrier18_Faults_0" bit 11
   1165: 'Carrier 18 Encoder Position Fault', class No Acknowledgement, trigger "DB302_HMI_Faults_Carrier18_Faults_0" bit 12
   1166: 'Carrier 18 Encoder Internal Error', class No Acknowledgement, trigger "DB302_HMI_Faults_Carrier18_Faults_0" bit 13
   1167: 'Carrier 18 Encoder Comm Fault', class No Acknowledgement, trigger "DB302_HMI_Faults_Carrier18_Faults_0" bit 14
   1168: 'Carrier 18 HMI Comm Fault', class No Acknowledgement, trigger "DB302_HMI_Faults_Carrier18_Faults_0" bit 15
   1169: 'Carrier 18 Crash Detection Fault', class No Acknowledgement, trigger "DB302_HMI_Faults_Carrier18_Faults_1" bit 0
   1170: 'Carrier 18 Carrier Number Invalid', class No Acknowledgement, trigger "DB302_HMI_Faults_Carrier18_Faults_1" bit 1
   1171: 'Carrier 18 Drive: PROFINET configuration error', class No Acknowledgement, trigger "DB302_HMI_Faults_Carrier18_Faults_1" bit 2
   1172: 'Carrier 18 Drive: Error internal communications', class No Acknowledgement, trigger "DB302_HMI_Faults_Carrier18_Faults_1" bit 3
   1173: 'Carrier 18 Drive: Motor overtemperature', class No Acknowledgement, trigger "DB302_HMI_Faults_Carrier18_Faults_1" bit 4
   1174: 'Carrier 18 Drive: Motor overcurrent', class No Acknowledgement, trigger "DB302_HMI_Faults_Carrier18_Faults_1" bit 5
   1175: 'Carrier 18 Drive: Infeed or power unit not ready', class No Acknowledgement, trigger "DB302_HMI_Faults_Carrier18_Faults_1" bit 6
   1176: 'Carrier 18 Drive: Short-circuit/ground fault detected', class No Acknowledgement, trigger "DB302_HMI_Faults_Carrier18_Faults_1" bit 7
   1177: 'Carrier 18 Drive: PROFINET Setpoint timeout', class No Acknowledgement, trigger "DB302_HMI_Faults_Carrier18_Faults_1" bit 8
   1178: 'Carrier 18 Power unit: Overcurrent', class No Acknowledgement, trigger "DB302_HMI_Faults_Carrier18_Faults_1" bit 9
   1179: 'Carrier 18 Power unit: DC link voltage overvoltage', class No Acknowledgement, trigger "DB302_HMI_Faults_Carrier18_Faults_1" bit 10
   1180: 'Carrier 18 Power unit: DC link voltage undervoltage', class No Acknowledgement, trigger "DB302_HMI_Faults_Carrier18_Faults_1" bit 11
   1181: 'Carrier 18 Power unit: Line phase failure in main circuit', class No Acknowledgement, trigger "DB302_HMI_Faults_Carrier18_Faults_1" bit 12
   1182: 'Carrier 18 Power unit: Phase failure motor cable', class No Acknowledgement, trigger "DB302_HMI_Faults_Carrier18_Faults_1" bit 13
   1183: 'Carrier 18 Power unit: Ground fault', class No Acknowledgement, trigger "DB302_HMI_Faults_Carrier18_Faults_1" bit 14
   1184: 'Spare_Fault_1184', class No Acknowledgement, trigger "DB302_HMI_Faults_Carrier18_Faults_1" bit 15
   1185: 'Carrier 18 Motion Off Fault', class No Acknowledgement, trigger "DB302_HMI_Faults_Carrier18_Faults_2" bit 0
   1186: 'Carrier 18 Motion On Fault', class No Acknowledgement, trigger "DB302_HMI_Faults_Carrier18_Faults_2" bit 1
   1187: 'Carrier 18 Spacing Fault', class No Acknowledgement, trigger "DB302_HMI_Faults_Carrier18_Faults_2" bit 2
   1188: 'Carrier 18 Duplicate Carrier Number Fault', class No Acknowledgement, trigger "DB302_HMI_Faults_Carrier18_Faults_2" bit 3
   1189: 'Spare_Fault_1189', class No Acknowledgement, trigger "DB302_HMI_Faults_Carrier18_Faults_2" bit 4
   1190: 'Spare_Fault_1190', class No Acknowledgement, trigger "DB302_HMI_Faults_Carrier18_Faults_2" bit 5
   1191: 'Spare_Fault_1191', class No Acknowledgement, trigger "DB302_HMI_Faults_Carrier18_Faults_2" bit 6
   1192: 'Spare_Fault_1192', class No Acknowledgement, trigger "DB302_HMI_Faults_Carrier18_Faults_2" bit 7
   1193: 'Spare_Fault_1193', class No Acknowledgement, trigger "DB302_HMI_Faults_Carrier18_Faults_2" bit 8
   1194: 'Spare_Fault_1194', class No Acknowledgement, trigger "DB302_HMI_Faults_Carrier18_Faults_2" bit 9
   1195: 'Spare_Fault_1195', class No Acknowledgement, trigger "DB302_HMI_Faults_Carrier18_Faults_2" bit 10
   1196: 'Spare_Fault_1196', class No Acknowledgement, trigger "DB302_HMI_Faults_Carrier18_Faults_2" bit 11
   1197: 'Spare_Fault_1197', class No Acknowledgement, trigger "DB302_HMI_Faults_Carrier18_Faults_2" bit 12
   1198: 'Spare_Fault_1198', class No Acknowledgement, trigger "DB302_HMI_Faults_Carrier18_Faults_2" bit 13
   1199: 'Spare_Fault_1199', class No Acknowledgement, trigger "DB302_HMI_Faults_Carrier18_Faults_2" bit 14
   1200: 'Spare_Fault_1200', class No Acknowledgement, trigger "DB302_HMI_Faults_Carrier18_Faults_2" bit 15
   1201: 'Spare_Fault_1201', class No Acknowledgement, trigger "DB302_HMI_Faults_Carrier18_Faults_3" bit 0
   1202: 'Spare_Fault_1202', class No Acknowledgement, trigger "DB302_HMI_Faults_Carrier18_Faults_3" bit 1
   1203: 'Spare_Fault_1203', class No Acknowledgement, trigger "DB302_HMI_Faults_Carrier18_Faults_3" bit 2
   1204: 'Spare_Fault_1204', class No Acknowledgement, trigger "DB302_HMI_Faults_Carrier18_Faults_3" bit 3
   1205: 'Spare_Fault_1205', class No Acknowledgement, trigger "DB302_HMI_Faults_Carrier18_Faults_3" bit 4
   1206: 'Spare_Fault_1206', class No Acknowledgement, trigger "DB302_HMI_Faults_Carrier18_Faults_3" bit 5
   1207: 'Spare_Fault_1207', class No Acknowledgement, trigger "DB302_HMI_Faults_Carrier18_Faults_3" bit 6
   1208: 'Spare_Fault_1208', class No Acknowledgement, trigger "DB302_HMI_Faults_Carrier18_Faults_3" bit 7
   1209: 'Spare_Fault_1209', class No Acknowledgement, trigger "DB302_HMI_Faults_Carrier18_Faults_3" bit 8
   1210: 'Spare_Fault_1210', class No Acknowledgement, trigger "DB302_HMI_Faults_Carrier18_Faults_3" bit 9
   1211: 'Spare_Fault_1211', class No Acknowledgement, trigger "DB302_HMI_Faults_Carrier18_Faults_3" bit 10
   1212: 'Spare_Fault_1212', class No Acknowledgement, trigger "DB302_HMI_Faults_Carrier18_Faults_3" bit 11
   1213: 'Spare_Fault_1213', class No Acknowledgement, trigger "DB302_HMI_Faults_Carrier18_Faults_3" bit 12
   1214: 'Spare_Fault_1214', class No Acknowledgement, trigger "DB302_HMI_Faults_Carrier18_Faults_3" bit 13
   1215: 'Spare_Fault_1215', class No Acknowledgement, trigger "DB302_HMI_Faults_Carrier18_Faults_3" bit 14
   1216: 'Spare_Fault_1216', class No Acknowledgement, trigger "DB302_HMI_Faults_Carrier18_Faults_3" bit 15
   1217: 'Carrier 19 Disconnect Open Power Fault DI11.0', class No Acknowledgement, trigger "DB302_HMI_Faults_Carrier19_Faults_0" bit 0
   1218: 'Carrier 19 Drive Profinet Comm Fault', class No Acknowledgement, trigger "DB302_HMI_Faults_Carrier19_Faults_0" bit 1
   1219: 'Carrier 19 Production Stop Not Reset', class No Acknowledgement, trigger "DB302_HMI_Faults_Carrier19_Faults_0" bit 2
   1220: 'Carrier 19 CB02122 Tripped', class No Acknowledgement, trigger "DB302_HMI_Faults_Carrier19_Faults_0" bit 3
   1221: 'Carrier 19 CB02123 Tripped', class No Acknowledgement, trigger "DB302_HMI_Faults_Carrier19_Faults_0" bit 4
   1222: 'Carrier 19 AUX1 CB Tripped', class No Acknowledgement, trigger "DB302_HMI_Faults_Carrier19_Faults_0" bit 5
   1223: 'Carrier 19 AUX2 CB Tripped', class No Acknowledgement, trigger "DB302_HMI_Faults_Carrier19_Faults_0" bit 6
   1224: 'Carrier 19 PLC Not Communicating', class No Acknowledgement, trigger "DB302_HMI_Faults_Carrier19_Faults_0" bit 7
   1225: 'Carrier 19 Safe Input Card Fault', class No Acknowledgement, trigger "DB302_HMI_Faults_Carrier19_Faults_0" bit 8
   1226: 'Carrier 19 Safe Output Card Fault', class No Acknowledgement, trigger "DB302_HMI_Faults_Carrier19_Faults_0" bit 9
   1227: 'Carrier 19 Standard Input Card Fault', class No Acknowledgement, trigger "DB302_HMI_Faults_Carrier19_Faults_0" bit 10
   1228: 'Carrier 19 Standard Output Card Fault', class No Acknowledgement, trigger "DB302_HMI_Faults_Carrier19_Faults_0" bit 11
   1229: 'Carrier 19 Encoder Position Fault', class No Acknowledgement, trigger "DB302_HMI_Faults_Carrier19_Faults_0" bit 12
   1230: 'Carrier 19 Encoder Internal Error', class No Acknowledgement, trigger "DB302_HMI_Faults_Carrier19_Faults_0" bit 13
   1231: 'Carrier 19 Encoder Comm Fault', class No Acknowledgement, trigger "DB302_HMI_Faults_Carrier19_Faults_0" bit 14
   1232: 'Carrier 19 HMI Comm Fault', class No Acknowledgement, trigger "DB302_HMI_Faults_Carrier19_Faults_0" bit 15
   1233: 'Carrier 19 Crash Detection Fault', class No Acknowledgement, trigger "DB302_HMI_Faults_Carrier19_Faults_1" bit 0
   1234: 'Carrier 19 Carrier Number Invalid', class No Acknowledgement, trigger "DB302_HMI_Faults_Carrier19_Faults_1" bit 1
   1235: 'Carrier 19 Drive: PROFINET configuration error', class No Acknowledgement, trigger "DB302_HMI_Faults_Carrier19_Faults_1" bit 2
   1236: 'Carrier 19 Drive: Error internal communications', class No Acknowledgement, trigger "DB302_HMI_Faults_Carrier19_Faults_1" bit 3
   1237: 'Carrier 19 Drive: Motor overtemperature', class No Acknowledgement, trigger "DB302_HMI_Faults_Carrier19_Faults_1" bit 4
   1238: 'Carrier 19 Drive: Motor overcurrent', class No Acknowledgement, trigger "DB302_HMI_Faults_Carrier19_Faults_1" bit 5
   1239: 'Carrier 19 Drive: Infeed or power unit not ready', class No Acknowledgement, trigger "DB302_HMI_Faults_Carrier19_Faults_1" bit 6
   1240: 'Carrier 19 Drive: Short-circuit/ground fault detected', class No Acknowledgement, trigger "DB302_HMI_Faults_Carrier19_Faults_1" bit 7
   1241: 'Carrier 19 Drive: PROFINET Setpoint timeout', class No Acknowledgement, trigger "DB302_HMI_Faults_Carrier19_Faults_1" bit 8
   1242: 'Carrier 19 Power unit: Overcurrent', class No Acknowledgement, trigger "DB302_HMI_Faults_Carrier19_Faults_1" bit 9
   1243: 'Carrier 19 Power unit: DC link voltage overvoltage', class No Acknowledgement, trigger "DB302_HMI_Faults_Carrier19_Faults_1" bit 10
   1244: 'Carrier 19 Power unit: DC link voltage undervoltage', class No Acknowledgement, trigger "DB302_HMI_Faults_Carrier19_Faults_1" bit 11
   1245: 'Carrier 19 Power unit: Line phase failure in main circuit', class No Acknowledgement, trigger "DB302_HMI_Faults_Carrier19_Faults_1" bit 12
   1246: 'Carrier 19 Power unit: Phase failure motor cable', class No Acknowledgement, trigger "DB302_HMI_Faults_Carrier19_Faults_1" bit 13
   1247: 'Carrier 19 Power unit: Ground fault', class No Acknowledgement, trigger "DB302_HMI_Faults_Carrier19_Faults_1" bit 14
   1248: 'Spare_Fault_1248', class No Acknowledgement, trigger "DB302_HMI_Faults_Carrier19_Faults_1" bit 15
   1249: 'Carrier 19 Motion Off Fault', class No Acknowledgement, trigger "DB302_HMI_Faults_Carrier19_Faults_2" bit 0
   1250: 'Carrier 19 Motion On Fault', class No Acknowledgement, trigger "DB302_HMI_Faults_Carrier19_Faults_2" bit 1
   1251: 'Carrier 19 Spacing Fault', class No Acknowledgement, trigger "DB302_HMI_Faults_Carrier19_Faults_2" bit 2
   1252: 'Carrier 19 Duplicate Carrier Number Fault', class No Acknowledgement, trigger "DB302_HMI_Faults_Carrier19_Faults_2" bit 3
   1253: 'Spare_Fault_1253', class No Acknowledgement, trigger "DB302_HMI_Faults_Carrier19_Faults_2" bit 4
   1254: 'Spare_Fault_1254', class No Acknowledgement, trigger "DB302_HMI_Faults_Carrier19_Faults_2" bit 5
   1255: 'Spare_Fault_1255', class No Acknowledgement, trigger "DB302_HMI_Faults_Carrier19_Faults_2" bit 6
   1256: 'Spare_Fault_1256', class No Acknowledgement, trigger "DB302_HMI_Faults_Carrier19_Faults_2" bit 7
   1257: 'Spare_Fault_1257', class No Acknowledgement, trigger "DB302_HMI_Faults_Carrier19_Faults_2" bit 8
   1258: 'Spare_Fault_1258', class No Acknowledgement, trigger "DB302_HMI_Faults_Carrier19_Faults_2" bit 9
   1259: 'Spare_Fault_1259', class No Acknowledgement, trigger "DB302_HMI_Faults_Carrier19_Faults_2" bit 10
   1260: 'Spare_Fault_1260', class No Acknowledgement, trigger "DB302_HMI_Faults_Carrier19_Faults_2" bit 11
   1261: 'Spare_Fault_1261', class No Acknowledgement, trigger "DB302_HMI_Faults_Carrier19_Faults_2" bit 12
   1262: 'Spare_Fault_1262', class No Acknowledgement, trigger "DB302_HMI_Faults_Carrier19_Faults_2" bit 13
   1263: 'Spare_Fault_1263', class No Acknowledgement, trigger "DB302_HMI_Faults_Carrier19_Faults_2" bit 14
   1264: 'Spare_Fault_1264', class No Acknowledgement, trigger "DB302_HMI_Faults_Carrier19_Faults_2" bit 15
   1265: 'Spare_Fault_1265', class No Acknowledgement, trigger "DB302_HMI_Faults_Carrier19_Faults_3" bit 0
   1266: 'Spare_Fault_1266', class No Acknowledgement, trigger "DB302_HMI_Faults_Carrier19_Faults_3" bit 1
   1267: 'Spare_Fault_1267', class No Acknowledgement, trigger "DB302_HMI_Faults_Carrier19_Faults_3" bit 2
   1268: 'Spare_Fault_1268', class No Acknowledgement, trigger "DB302_HMI_Faults_Carrier19_Faults_3" bit 3
   1269: 'Spare_Fault_1269', class No Acknowledgement, trigger "DB302_HMI_Faults_Carrier19_Faults_3" bit 4
   1270: 'Spare_Fault_1270', class No Acknowledgement, trigger "DB302_HMI_Faults_Carrier19_Faults_3" bit 5
   1271: 'Spare_Fault_1271', class No Acknowledgement, trigger "DB302_HMI_Faults_Carrier19_Faults_3" bit 6
   1272: 'Spare_Fault_1272', class No Acknowledgement, trigger "DB302_HMI_Faults_Carrier19_Faults_3" bit 7
   1273: 'Spare_Fault_1273', class No Acknowledgement, trigger "DB302_HMI_Faults_Carrier19_Faults_3" bit 8
   1274: 'Spare_Fault_1274', class No Acknowledgement, trigger "DB302_HMI_Faults_Carrier19_Faults_3" bit 9
   1275: 'Spare_Fault_1275', class No Acknowledgement, trigger "DB302_HMI_Faults_Carrier19_Faults_3" bit 10
   1276: 'Spare_Fault_1276', class No Acknowledgement, trigger "DB302_HMI_Faults_Carrier19_Faults_3" bit 11
   1277: 'Spare_Fault_1277', class No Acknowledgement, trigger "DB302_HMI_Faults_Carrier19_Faults_3" bit 12
   1278: 'Spare_Fault_1278', class No Acknowledgement, trigger "DB302_HMI_Faults_Carrier19_Faults_3" bit 13
   1279: 'Spare_Fault_1279', class No Acknowledgement, trigger "DB302_HMI_Faults_Carrier19_Faults_3" bit 14
   1280: 'Spare_Fault_1280', class No Acknowledgement, trigger "DB302_HMI_Faults_Carrier19_Faults_3" bit 15
   1281: 'Carrier 20 Disconnect Open Power Fault DI11.0', class No Acknowledgement, trigger "DB302_HMI_Faults_Carrier20_Faults_0" bit 0
   1282: 'Carrier 20 Drive Profinet Comm Fault', class No Acknowledgement, trigger "DB302_HMI_Faults_Carrier20_Faults_0" bit 1
   1283: 'Carrier 20 Production Stop Not Reset', class No Acknowledgement, trigger "DB302_HMI_Faults_Carrier20_Faults_0" bit 2
   1284: 'Carrier 20 CB02122 Tripped', class No Acknowledgement, trigger "DB302_HMI_Faults_Carrier20_Faults_0" bit 3
   1285: 'Carrier 20 CB02123 Tripped', class No Acknowledgement, trigger "DB302_HMI_Faults_Carrier20_Faults_0" bit 4
   1286: 'Carrier 20 AUX1 CB Tripped', class No Acknowledgement, trigger "DB302_HMI_Faults_Carrier20_Faults_0" bit 5
   1287: 'Carrier 20 AUX2 CB Tripped', class No Acknowledgement, trigger "DB302_HMI_Faults_Carrier20_Faults_0" bit 6
   1288: 'Carrier 20 PLC Not Communicating', class No Acknowledgement, trigger "DB302_HMI_Faults_Carrier20_Faults_0" bit 7
   1289: 'Carrier 20 Safe Input Card Fault', class No Acknowledgement, trigger "DB302_HMI_Faults_Carrier20_Faults_0" bit 8